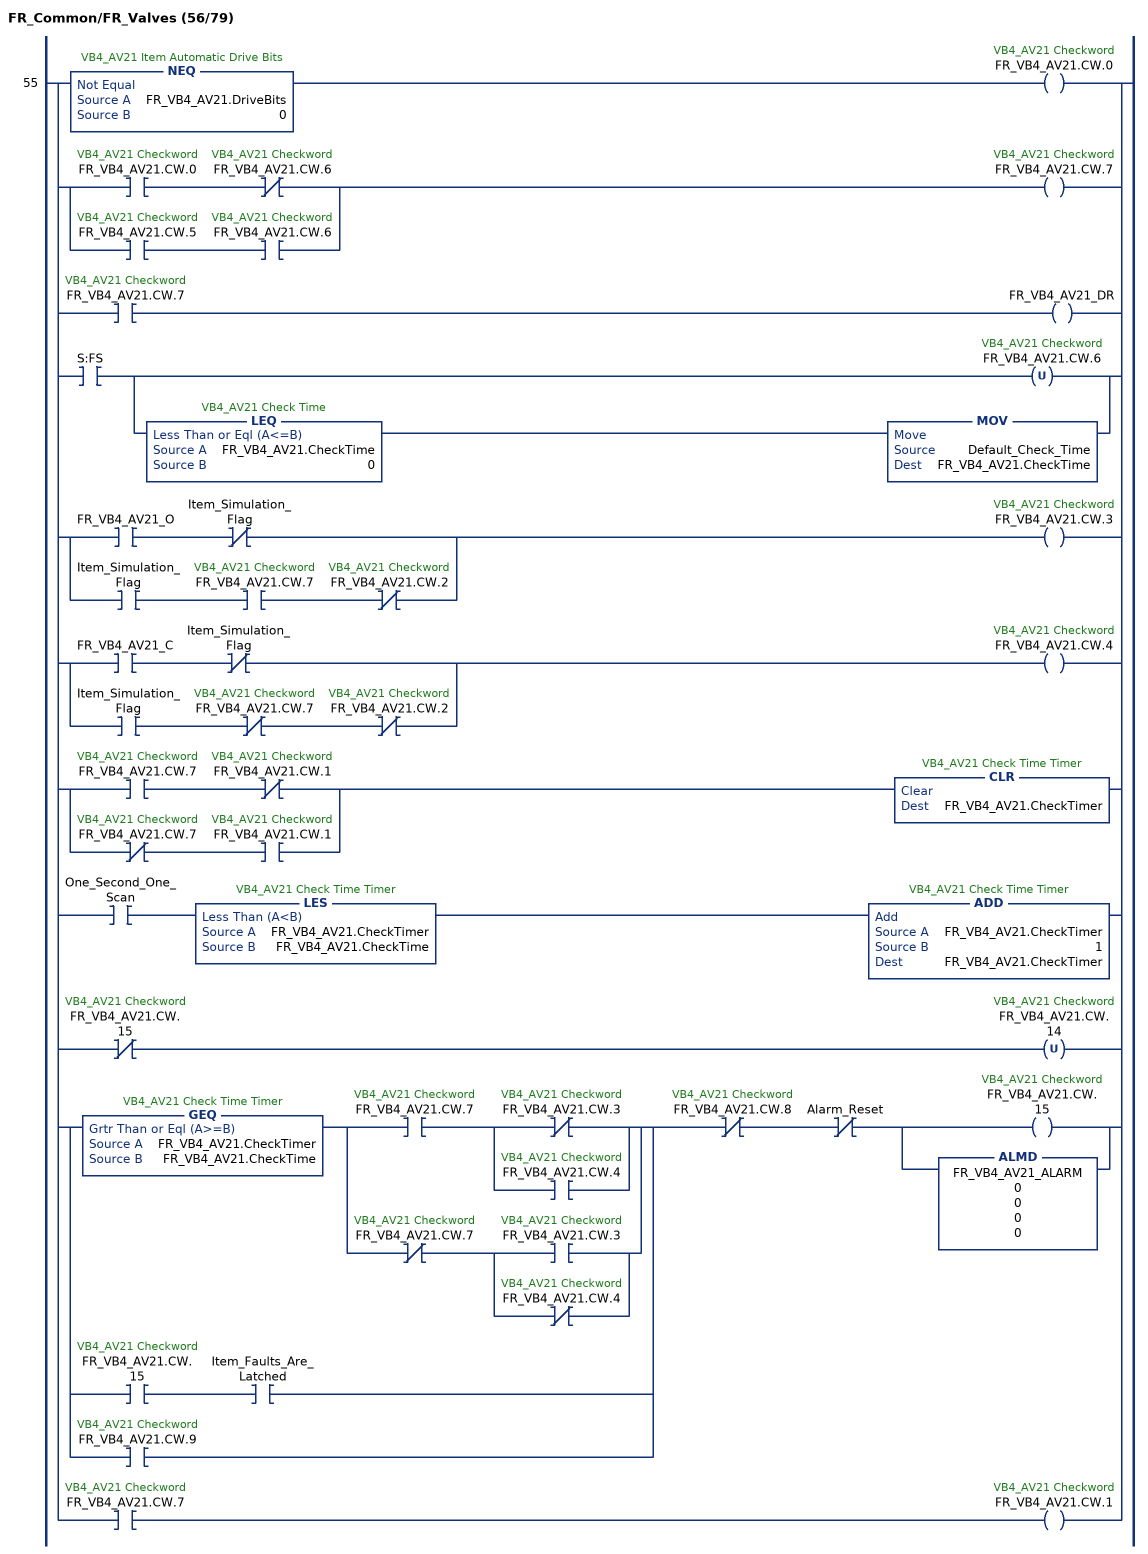
   55: [NEQ(FR_VB4_AV21.DriveBits,0) OTE(FR_VB4_AV21.CW.0) ,[XIC(FR_VB4_AV21.CW.0) XIO(FR_VB4_AV21.CW.6) ,XIC(FR_VB4_AV21.CW.5) XIC(FR_VB4_AV21.CW.6) ] OTE(FR_VB4_AV21.CW.7) ,XIC(FR_VB4_AV21.CW.7) OTE(FR_VB4_AV21_DR) ,XIC(S:FS) [OTU(FR_VB4_AV21.CW.6) ,LEQ(FR_VB4_AV21.CheckTime,0) MOV(Default_Check_Time,FR_VB4_AV21.CheckTime) ] ,[[XIC(FR_VB4_AV21_O) XIO(Item_Simulation_Flag) ,XIC(Item_Simulation_Flag) XIC(FR_VB4_AV21.CW.7) XIO(FR_VB4_AV21.CW.2) ] OTE(FR_VB4_AV21.CW.3) ,[XIC(FR_VB4_AV21_C) XIO(Item_Simulation_Flag) ,XIC(Item_Simulation_Flag) XIO(FR_VB4_AV21.CW.7) XIO(FR_VB4_AV21.CW.2) ] OTE(FR_VB4_AV21.CW.4) ] ,[XIC(FR_VB4_AV21.CW.7) XIO(FR_VB4_AV21.CW.1) ,XIO(FR_VB4_AV21.CW.7) XIC(FR_VB4_AV21.CW.1) ] CLR(FR_VB4_AV21.CheckTimer) ,XIC(One_Second_One_Scan) LES(FR_VB4_AV21.CheckTimer,FR_VB4_AV21.CheckTime) ADD(FR_VB4_AV21.CheckTimer,1,FR_VB4_AV21.CheckTimer) ,XIO(FR_VB4_AV21.CW.15) OTU(FR_VB4_AV21.CW.14) ,[GEQ(FR_VB4_AV21.CheckTimer,FR_VB4_AV21.CheckTime) [XIC(FR_VB4_AV21.CW.7) [XIO(FR_VB4_AV21.CW.3) ,XIC(FR_VB4_AV21.CW.4) ] ,XIO(FR_VB4_AV21.CW.7) [XIC(FR_VB4_AV21.CW.3) ,XIO(FR_VB4_AV21.CW.4) ] ] ,XIC(FR_VB4_AV21.CW.15) XIC(Item_Faults_Are_Latched) ,XIC(FR_VB4_AV21.CW.9) ] XIO(FR_VB4_AV21.CW.8) XIO(Alarm_Reset) [OTE(FR_VB4_AV21.CW.15) ,ALMD(FR_VB4_AV21_ALARM,0,0,0,0) ] ,XIC(FR_VB4_AV21.CW.7) OTE(FR_VB4_AV21.CW.1) ];
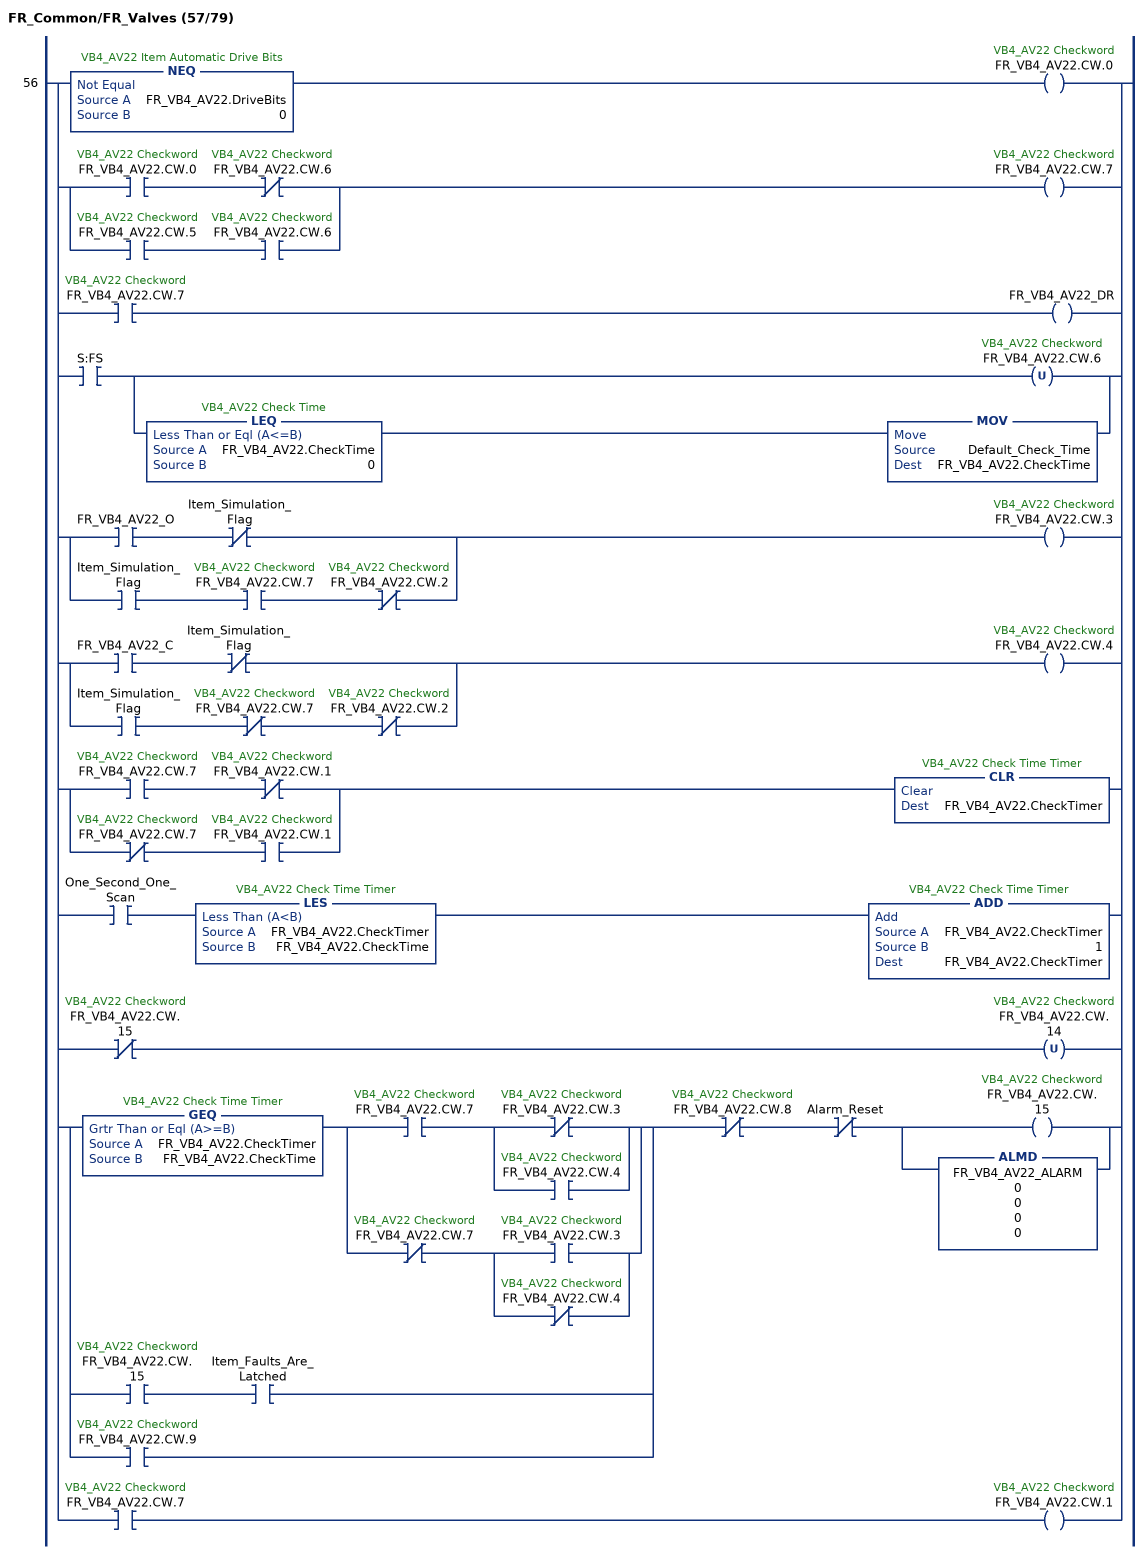
   56: [NEQ(FR_VB4_AV22.DriveBits,0) OTE(FR_VB4_AV22.CW.0) ,[XIC(FR_VB4_AV22.CW.0) XIO(FR_VB4_AV22.CW.6) ,XIC(FR_VB4_AV22.CW.5) XIC(FR_VB4_AV22.CW.6) ] OTE(FR_VB4_AV22.CW.7) ,XIC(FR_VB4_AV22.CW.7) OTE(FR_VB4_AV22_DR) ,XIC(S:FS) [OTU(FR_VB4_AV22.CW.6) ,LEQ(FR_VB4_AV22.CheckTime,0) MOV(Default_Check_Time,FR_VB4_AV22.CheckTime) ] ,[[XIC(FR_VB4_AV22_O) XIO(Item_Simulation_Flag) ,XIC(Item_Simulation_Flag) XIC(FR_VB4_AV22.CW.7) XIO(FR_VB4_AV22.CW.2) ] OTE(FR_VB4_AV22.CW.3) ,[XIC(FR_VB4_AV22_C) XIO(Item_Simulation_Flag) ,XIC(Item_Simulation_Flag) XIO(FR_VB4_AV22.CW.7) XIO(FR_VB4_AV22.CW.2) ] OTE(FR_VB4_AV22.CW.4) ] ,[XIC(FR_VB4_AV22.CW.7) XIO(FR_VB4_AV22.CW.1) ,XIO(FR_VB4_AV22.CW.7) XIC(FR_VB4_AV22.CW.1) ] CLR(FR_VB4_AV22.CheckTimer) ,XIC(One_Second_One_Scan) LES(FR_VB4_AV22.CheckTimer,FR_VB4_AV22.CheckTime) ADD(FR_VB4_AV22.CheckTimer,1,FR_VB4_AV22.CheckTimer) ,XIO(FR_VB4_AV22.CW.15) OTU(FR_VB4_AV22.CW.14) ,[GEQ(FR_VB4_AV22.CheckTimer,FR_VB4_AV22.CheckTime) [XIC(FR_VB4_AV22.CW.7) [XIO(FR_VB4_AV22.CW.3) ,XIC(FR_VB4_AV22.CW.4) ] ,XIO(FR_VB4_AV22.CW.7) [XIC(FR_VB4_AV22.CW.3) ,XIO(FR_VB4_AV22.CW.4) ] ] ,XIC(FR_VB4_AV22.CW.15) XIC(Item_Faults_Are_Latched) ,XIC(FR_VB4_AV22.CW.9) ] XIO(FR_VB4_AV22.CW.8) XIO(Alarm_Reset) [OTE(FR_VB4_AV22.CW.15) ,ALMD(FR_VB4_AV22_ALARM,0,0,0,0) ] ,XIC(FR_VB4_AV22.CW.7) OTE(FR_VB4_AV22.CW.1) ];
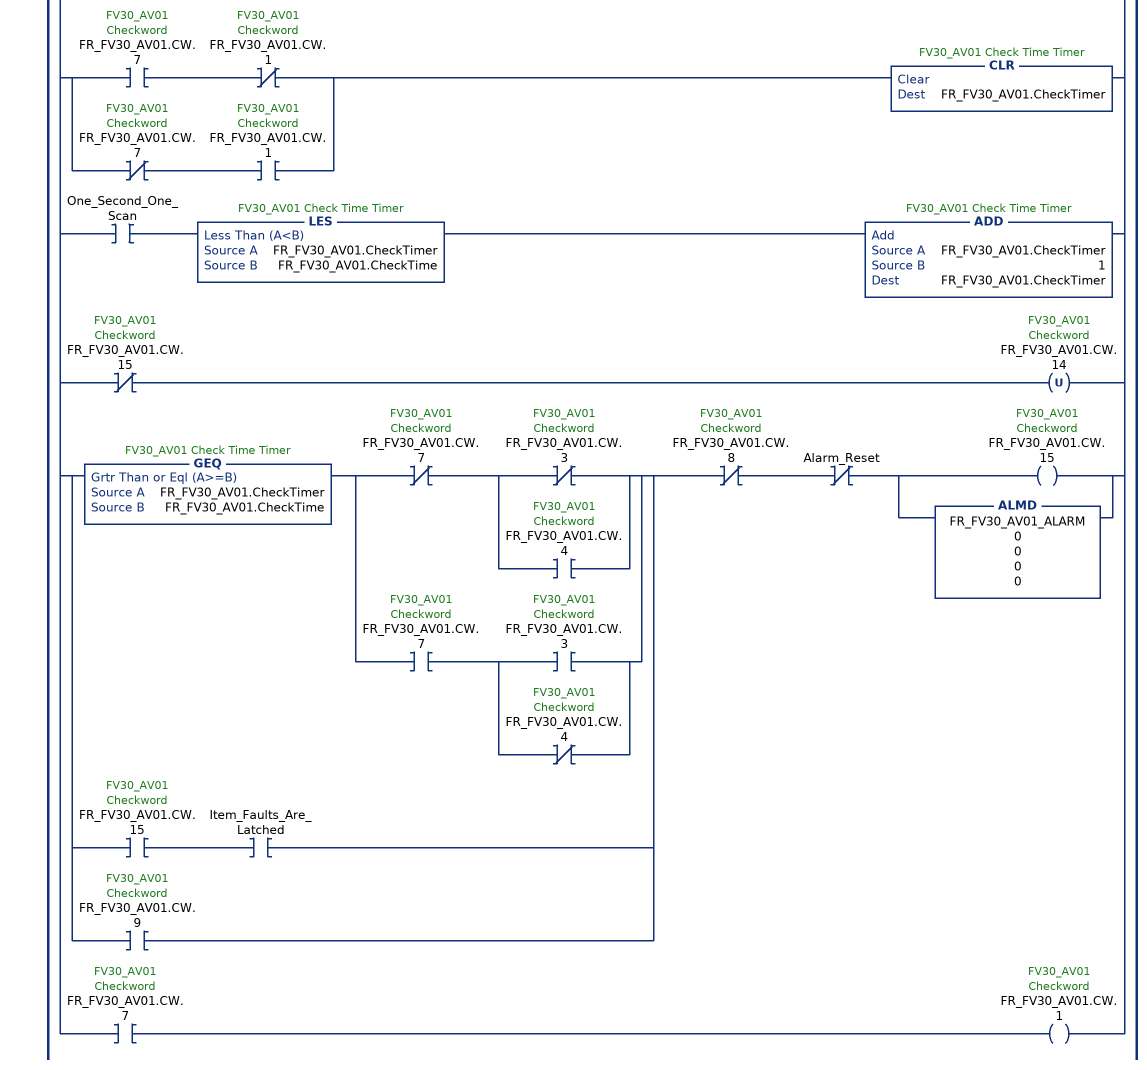
   57: [NEQ(FR_FV30_AV01.DriveBits,0) OTE(FR_FV30_AV01.CW.0) ,[XIC(FR_FV30_AV01.CW.0) XIO(FR_FV30_AV01.CW.6) ,XIC(FR_FV30_AV01.CW.5) XIC(FR_FV30_AV01.CW.6) ] OTE(FR_FV30_AV01.CW.7) ,XIC(FR_FV30_AV01.CW.7) OTE(FR_FV30_AV01_RDR) ,XIC(S:FS) [OTU(FR_FV30_AV01.CW.6) ,LEQ(FR_FV30_AV01.CheckTime,0) MOV(Default_Check_Time,FR_FV30_AV01.CheckTime) ] ,[[XIC(FR_FV30_AV01_O) XIO(Item_Simulation_Flag) ,XIC(Item_Simulation_Flag) XIO(FR_FV30_AV01.CW.7) XIO(FR_FV30_AV01.CW.2) ] OTE(FR_FV30_AV01.CW.3) ,[XIC(FR_FV30_AV01_C) XIO(Item_Simulation_Flag) ,XIC(Item_Simulation_Flag) XIC(FR_FV30_AV01.CW.7) XIO(FR_FV30_AV01.CW.2) ] OTE(FR_FV30_AV01.CW.4) ] ,[XIC(FR_FV30_AV01.CW.7) XIO(FR_FV30_AV01.CW.1) ,XIO(FR_FV30_AV01.CW.7) XIC(FR_FV30_AV01.CW.1) ] CLR(FR_FV30_AV01.CheckTimer) ,XIC(One_Second_One_Scan) LES(FR_FV30_AV01.CheckTimer,FR_FV30_AV01.CheckTime) ADD(FR_FV30_AV01.CheckTimer,1,FR_FV30_AV01.CheckTimer) ,XIO(FR_FV30_AV01.CW.15) OTU(FR_FV30_AV01.CW.14) ,[GEQ(FR_FV30_AV01.CheckTimer,FR_FV30_AV01.CheckTime) [XIO(FR_FV30_AV01.CW.7) [XIO(FR_FV30_AV01.CW.3) ,XIC(FR_FV30_AV01.CW.4) ] ,XIC(FR_FV30_AV01.CW.7) [XIC(FR_FV30_AV01.CW.3) ,XIO(FR_FV30_AV01.CW.4) ] ] ,XIC(FR_FV30_AV01.CW.15) XIC(Item_Faults_Are_Latched) ,XIC(FR_FV30_AV01.CW.9) ] XIO(FR_FV30_AV01.CW.8) XIO(Alarm_Reset) [OTE(FR_FV30_AV01.CW.15) ,ALMD(FR_FV30_AV01_ALARM,0,0,0,0) ] ,XIC(FR_FV30_AV01.CW.7) OTE(FR_FV30_AV01.CW.1) ];
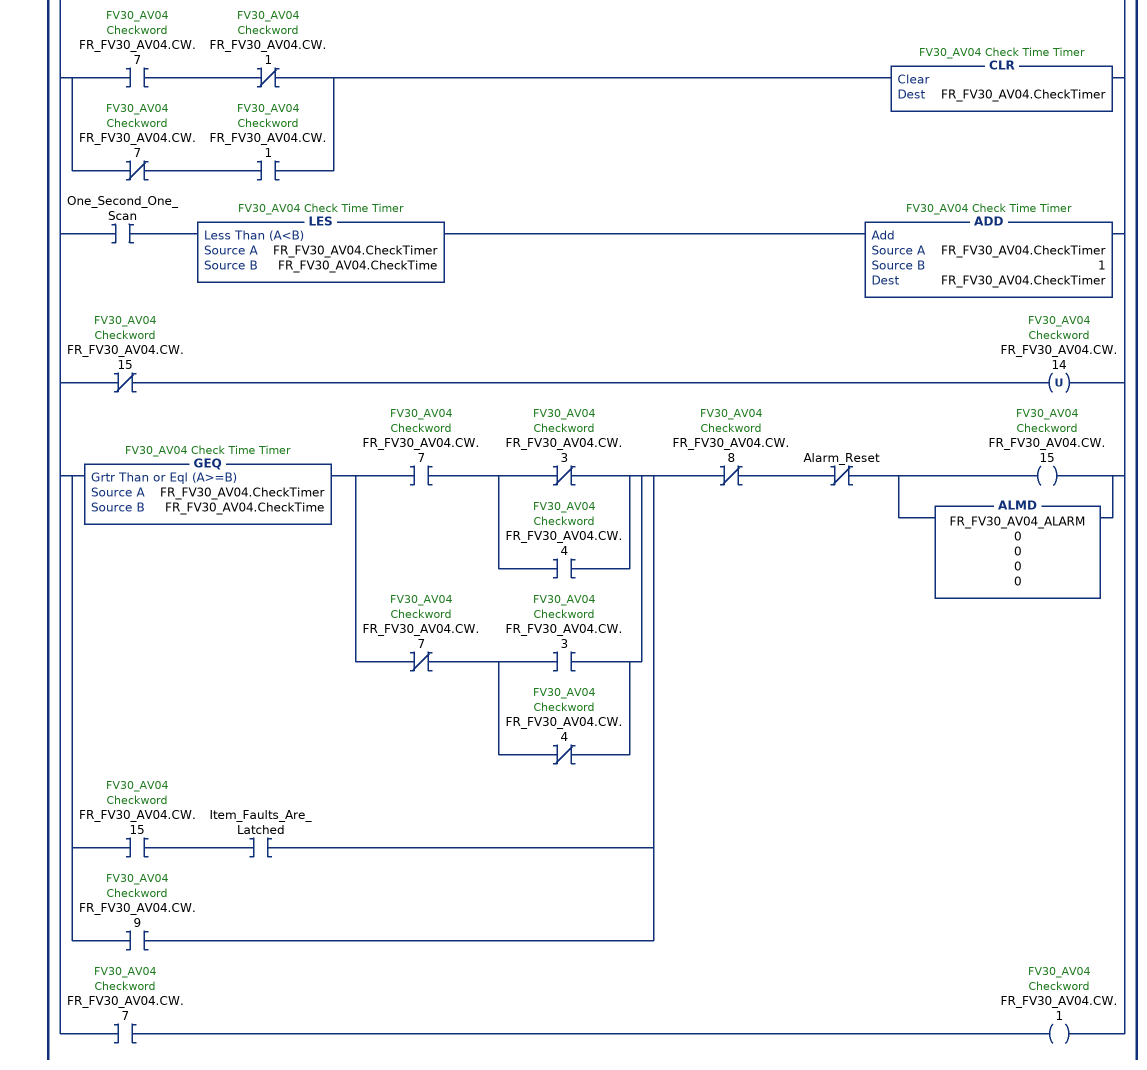
   58: [NEQ(FR_FV30_AV04.DriveBits,0) OTE(FR_FV30_AV04.CW.0) ,[XIC(FR_FV30_AV04.CW.0) XIO(FR_FV30_AV04.CW.6) ,XIC(FR_FV30_AV04.CW.5) XIC(FR_FV30_AV04.CW.6) ] OTE(FR_FV30_AV04.CW.7) ,XIC(FR_FV30_AV04.CW.7) OTE(FR_FV30_AV04_DR) ,XIC(S:FS) [OTU(FR_FV30_AV04.CW.6) ,LEQ(FR_FV30_AV04.CheckTime,0) MOV(Default_Check_Time,FR_FV30_AV04.CheckTime) ] ,[[XIC(FR_FV30_AV04_O) XIO(Item_Simulation_Flag) ,XIC(Item_Simulation_Flag) XIC(FR_FV30_AV04.CW.7) XIO(FR_FV30_AV04.CW.2) ] OTE(FR_FV30_AV04.CW.3) ,[XIC(FR_FV30_AV04_C) XIO(Item_Simulation_Flag) ,XIC(Item_Simulation_Flag) XIO(FR_FV30_AV04.CW.7) XIO(FR_FV30_AV04.CW.2) ] OTE(FR_FV30_AV04.CW.4) ] ,[XIC(FR_FV30_AV04.CW.7) XIO(FR_FV30_AV04.CW.1) ,XIO(FR_FV30_AV04.CW.7) XIC(FR_FV30_AV04.CW.1) ] CLR(FR_FV30_AV04.CheckTimer) ,XIC(One_Second_One_Scan) LES(FR_FV30_AV04.CheckTimer,FR_FV30_AV04.CheckTime) ADD(FR_FV30_AV04.CheckTimer,1,FR_FV30_AV04.CheckTimer) ,XIO(FR_FV30_AV04.CW.15) OTU(FR_FV30_AV04.CW.14) ,[GEQ(FR_FV30_AV04.CheckTimer,FR_FV30_AV04.CheckTime) [XIC(FR_FV30_AV04.CW.7) [XIO(FR_FV30_AV04.CW.3) ,XIC(FR_FV30_AV04.CW.4) ] ,XIO(FR_FV30_AV04.CW.7) [XIC(FR_FV30_AV04.CW.3) ,XIO(FR_FV30_AV04.CW.4) ] ] ,XIC(FR_FV30_AV04.CW.15) XIC(Item_Faults_Are_Latched) ,XIC(FR_FV30_AV04.CW.9) ] XIO(FR_FV30_AV04.CW.8) XIO(Alarm_Reset) [OTE(FR_FV30_AV04.CW.15) ,ALMD(FR_FV30_AV04_ALARM,0,0,0,0) ] ,XIC(FR_FV30_AV04.CW.7) OTE(FR_FV30_AV04.CW.1) ];
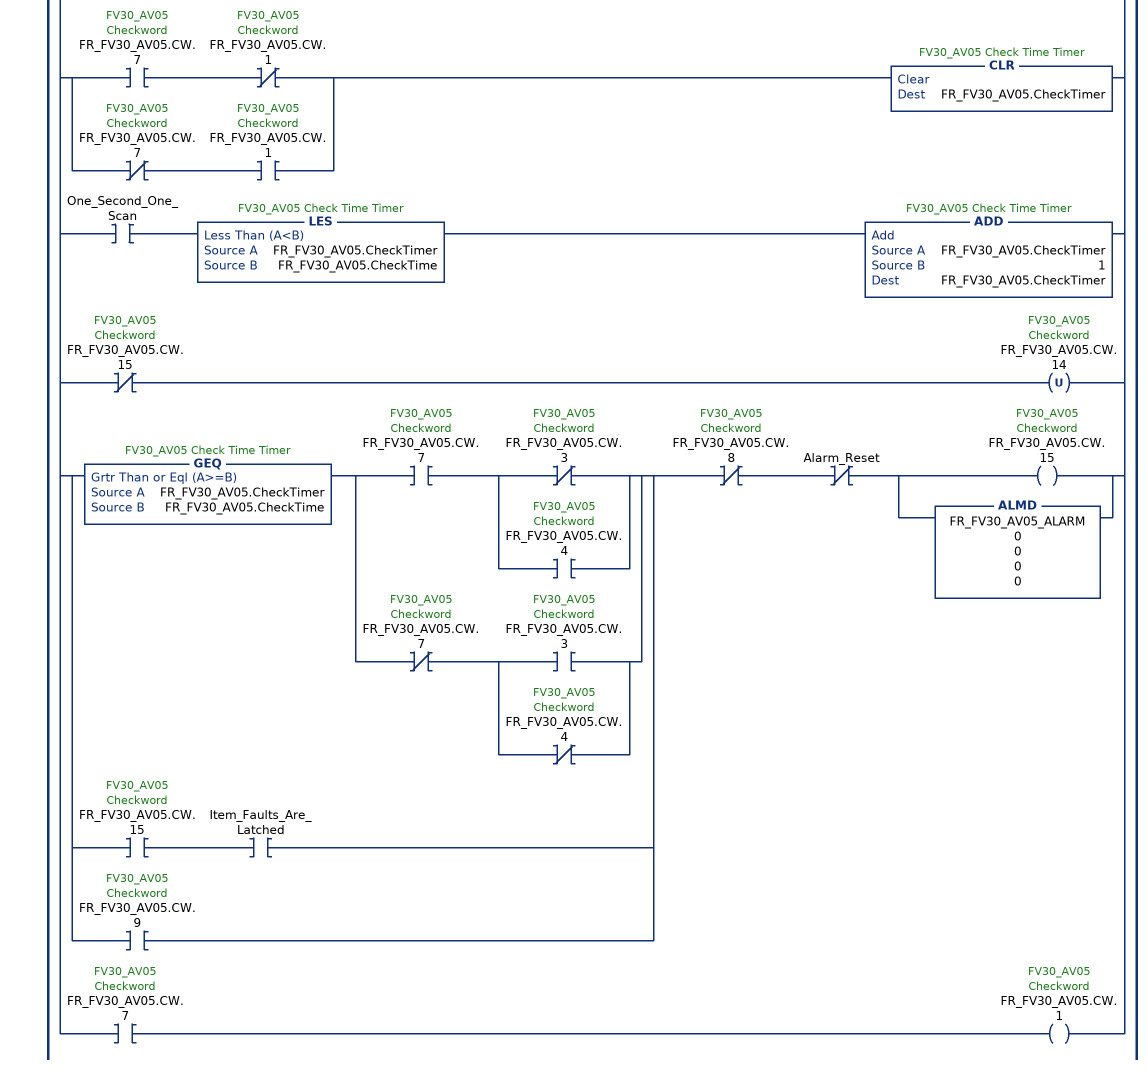
   59: [NEQ(FR_FV30_AV05.DriveBits,0) OTE(FR_FV30_AV05.CW.0) ,[XIC(FR_FV30_AV05.CW.0) XIO(FR_FV30_AV05.CW.6) ,XIC(FR_FV30_AV05.CW.5) XIC(FR_FV30_AV05.CW.6) ] OTE(FR_FV30_AV05.CW.7) ,XIC(FR_FV30_AV05.CW.7) OTE(FR_FV30_AV05_DR) ,XIC(S:FS) [OTU(FR_FV30_AV05.CW.6) ,LEQ(FR_FV30_AV05.CheckTime,0) MOV(Default_Check_Time,FR_FV30_AV05.CheckTime) ] ,[[XIC(FR_FV30_AV05_O) XIO(Item_Simulation_Flag) ,XIC(Item_Simulation_Flag) XIC(FR_FV30_AV05.CW.7) XIO(FR_FV30_AV05.CW.2) ] OTE(FR_FV30_AV05.CW.3) ,[XIC(FR_FV30_AV05_C) XIO(Item_Simulation_Flag) ,XIC(Item_Simulation_Flag) XIO(FR_FV30_AV05.CW.7) XIO(FR_FV30_AV05.CW.2) ] OTE(FR_FV30_AV05.CW.4) ] ,[XIC(FR_FV30_AV05.CW.7) XIO(FR_FV30_AV05.CW.1) ,XIO(FR_FV30_AV05.CW.7) XIC(FR_FV30_AV05.CW.1) ] CLR(FR_FV30_AV05.CheckTimer) ,XIC(One_Second_One_Scan) LES(FR_FV30_AV05.CheckTimer,FR_FV30_AV05.CheckTime) ADD(FR_FV30_AV05.CheckTimer,1,FR_FV30_AV05.CheckTimer) ,XIO(FR_FV30_AV05.CW.15) OTU(FR_FV30_AV05.CW.14) ,[GEQ(FR_FV30_AV05.CheckTimer,FR_FV30_AV05.CheckTime) [XIC(FR_FV30_AV05.CW.7) [XIO(FR_FV30_AV05.CW.3) ,XIC(FR_FV30_AV05.CW.4) ] ,XIO(FR_FV30_AV05.CW.7) [XIC(FR_FV30_AV05.CW.3) ,XIO(FR_FV30_AV05.CW.4) ] ] ,XIC(FR_FV30_AV05.CW.15) XIC(Item_Faults_Are_Latched) ,XIC(FR_FV30_AV05.CW.9) ] XIO(FR_FV30_AV05.CW.8) XIO(Alarm_Reset) [OTE(FR_FV30_AV05.CW.15) ,ALMD(FR_FV30_AV05_ALARM,0,0,0,0) ] ,XIC(FR_FV30_AV05.CW.7) OTE(FR_FV30_AV05.CW.1) ];
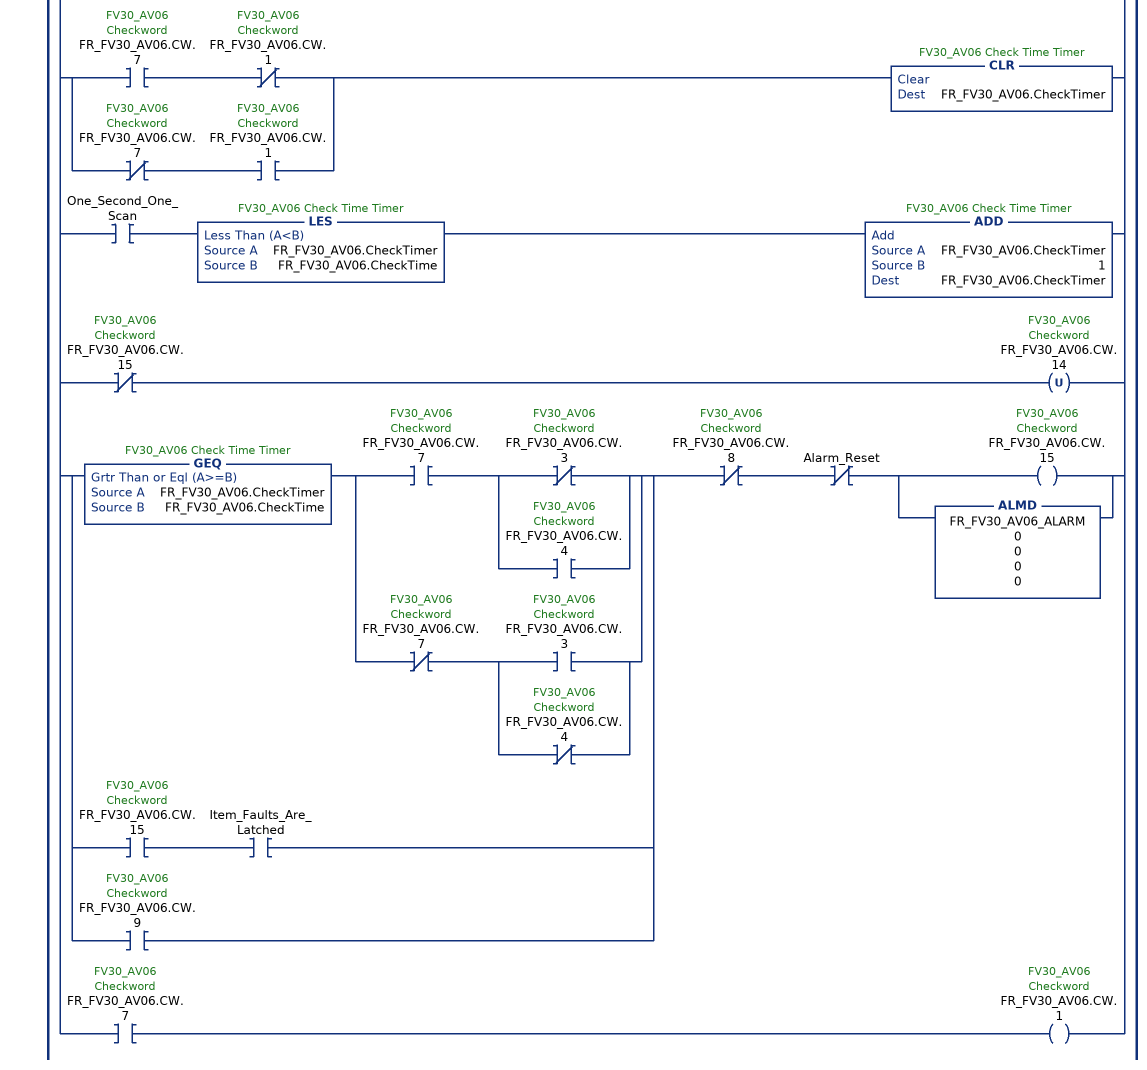
   60: [NEQ(FR_FV30_AV06.DriveBits,0) OTE(FR_FV30_AV06.CW.0) ,[XIC(FR_FV30_AV06.CW.0) XIO(FR_FV30_AV06.CW.6) ,XIC(FR_FV30_AV06.CW.5) XIC(FR_FV30_AV06.CW.6) ] OTE(FR_FV30_AV06.CW.7) ,XIC(FR_FV30_AV06.CW.7) OTE(FR_FV30_AV06_DR) ,XIC(S:FS) [OTU(FR_FV30_AV06.CW.6) ,LEQ(FR_FV30_AV06.CheckTime,0) MOV(Default_Check_Time,FR_FV30_AV06.CheckTime) ] ,[[XIC(FR_FV30_AV06_O) XIO(Item_Simulation_Flag) ,XIC(Item_Simulation_Flag) XIC(FR_FV30_AV06.CW.7) XIO(FR_FV30_AV06.CW.2) ] OTE(FR_FV30_AV06.CW.3) ,[XIC(FR_FV30_AV06_C) XIO(Item_Simulation_Flag) ,XIC(Item_Simulation_Flag) XIO(FR_FV30_AV06.CW.7) XIO(FR_FV30_AV06.CW.2) ] OTE(FR_FV30_AV06.CW.4) ] ,[XIC(FR_FV30_AV06.CW.7) XIO(FR_FV30_AV06.CW.1) ,XIO(FR_FV30_AV06.CW.7) XIC(FR_FV30_AV06.CW.1) ] CLR(FR_FV30_AV06.CheckTimer) ,XIC(One_Second_One_Scan) LES(FR_FV30_AV06.CheckTimer,FR_FV30_AV06.CheckTime) ADD(FR_FV30_AV06.CheckTimer,1,FR_FV30_AV06.CheckTimer) ,XIO(FR_FV30_AV06.CW.15) OTU(FR_FV30_AV06.CW.14) ,[GEQ(FR_FV30_AV06.CheckTimer,FR_FV30_AV06.CheckTime) [XIC(FR_FV30_AV06.CW.7) [XIO(FR_FV30_AV06.CW.3) ,XIC(FR_FV30_AV06.CW.4) ] ,XIO(FR_FV30_AV06.CW.7) [XIC(FR_FV30_AV06.CW.3) ,XIO(FR_FV30_AV06.CW.4) ] ] ,XIC(FR_FV30_AV06.CW.15) XIC(Item_Faults_Are_Latched) ,XIC(FR_FV30_AV06.CW.9) ] XIO(FR_FV30_AV06.CW.8) XIO(Alarm_Reset) [OTE(FR_FV30_AV06.CW.15) ,ALMD(FR_FV30_AV06_ALARM,0,0,0,0) ] ,XIC(FR_FV30_AV06.CW.7) OTE(FR_FV30_AV06.CW.1) ];
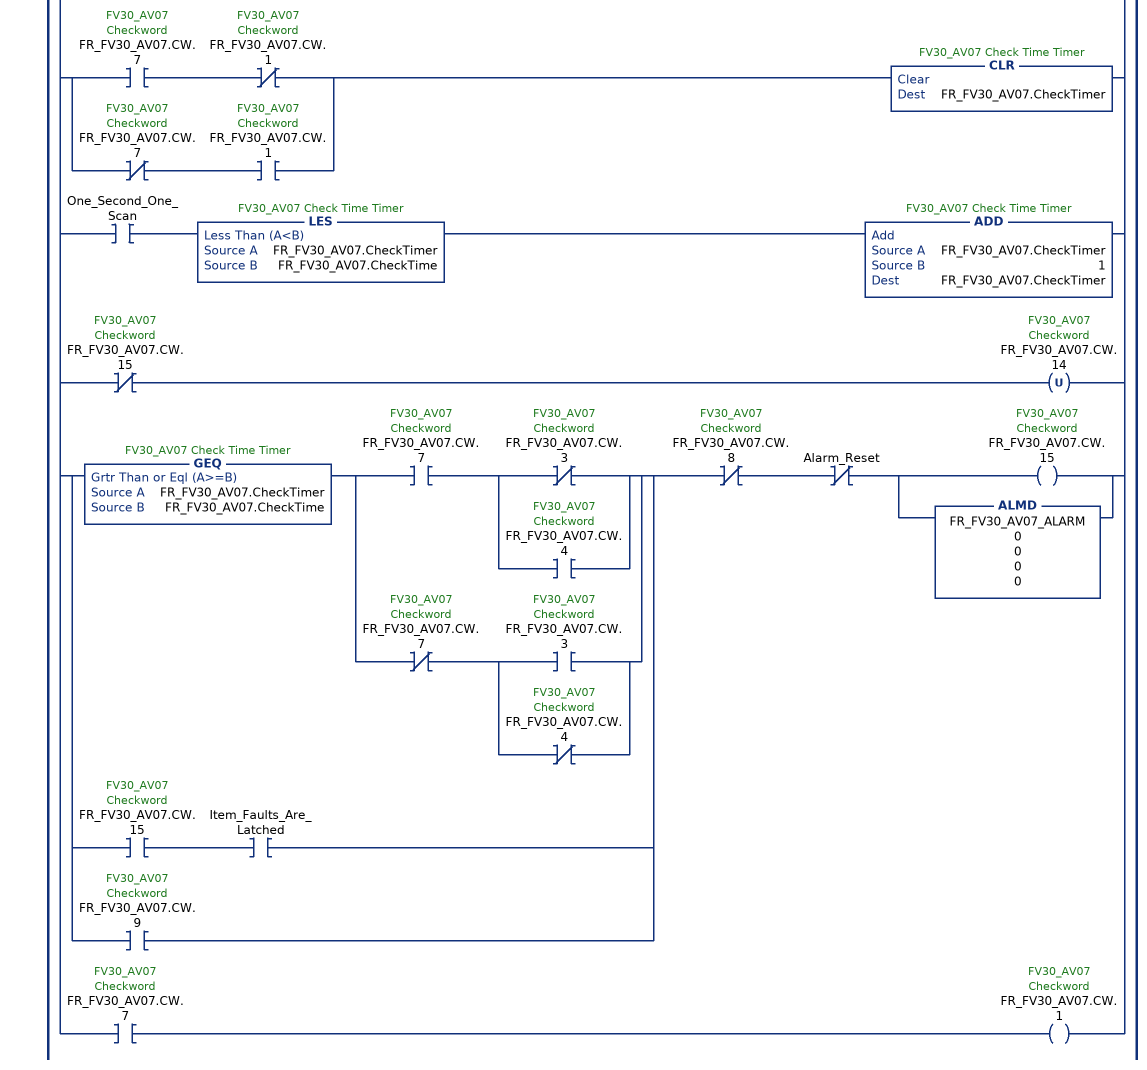
   61: [NEQ(FR_FV30_AV07.DriveBits,0) OTE(FR_FV30_AV07.CW.0) ,[XIC(FR_FV30_AV07.CW.0) XIO(FR_FV30_AV07.CW.6) ,XIC(FR_FV30_AV07.CW.5) XIC(FR_FV30_AV07.CW.6) ] OTE(FR_FV30_AV07.CW.7) ,XIC(FR_FV30_AV07.CW.7) OTE(FR_FV30_AV07_DR) ,XIC(S:FS) [OTU(FR_FV30_AV07.CW.6) ,LEQ(FR_FV30_AV07.CheckTime,0) MOV(Default_Check_Time,FR_FV30_AV07.CheckTime) ] ,[[XIC(FR_FV30_AV07_O) XIO(Item_Simulation_Flag) ,XIC(Item_Simulation_Flag) XIC(FR_FV30_AV07.CW.7) XIO(FR_FV30_AV07.CW.2) ] OTE(FR_FV30_AV07.CW.3) ,[XIC(FR_FV30_AV07_C) XIO(Item_Simulation_Flag) ,XIC(Item_Simulation_Flag) XIO(FR_FV30_AV07.CW.7) XIO(FR_FV30_AV07.CW.2) ] OTE(FR_FV30_AV07.CW.4) ] ,[XIC(FR_FV30_AV07.CW.7) XIO(FR_FV30_AV07.CW.1) ,XIO(FR_FV30_AV07.CW.7) XIC(FR_FV30_AV07.CW.1) ] CLR(FR_FV30_AV07.CheckTimer) ,XIC(One_Second_One_Scan) LES(FR_FV30_AV07.CheckTimer,FR_FV30_AV07.CheckTime) ADD(FR_FV30_AV07.CheckTimer,1,FR_FV30_AV07.CheckTimer) ,XIO(FR_FV30_AV07.CW.15) OTU(FR_FV30_AV07.CW.14) ,[GEQ(FR_FV30_AV07.CheckTimer,FR_FV30_AV07.CheckTime) [XIC(FR_FV30_AV07.CW.7) [XIO(FR_FV30_AV07.CW.3) ,XIC(FR_FV30_AV07.CW.4) ] ,XIO(FR_FV30_AV07.CW.7) [XIC(FR_FV30_AV07.CW.3) ,XIO(FR_FV30_AV07.CW.4) ] ] ,XIC(FR_FV30_AV07.CW.15) XIC(Item_Faults_Are_Latched) ,XIC(FR_FV30_AV07.CW.9) ] XIO(FR_FV30_AV07.CW.8) XIO(Alarm_Reset) [OTE(FR_FV30_AV07.CW.15) ,ALMD(FR_FV30_AV07_ALARM,0,0,0,0) ] ,XIC(FR_FV30_AV07.CW.7) OTE(FR_FV30_AV07.CW.1) ];
